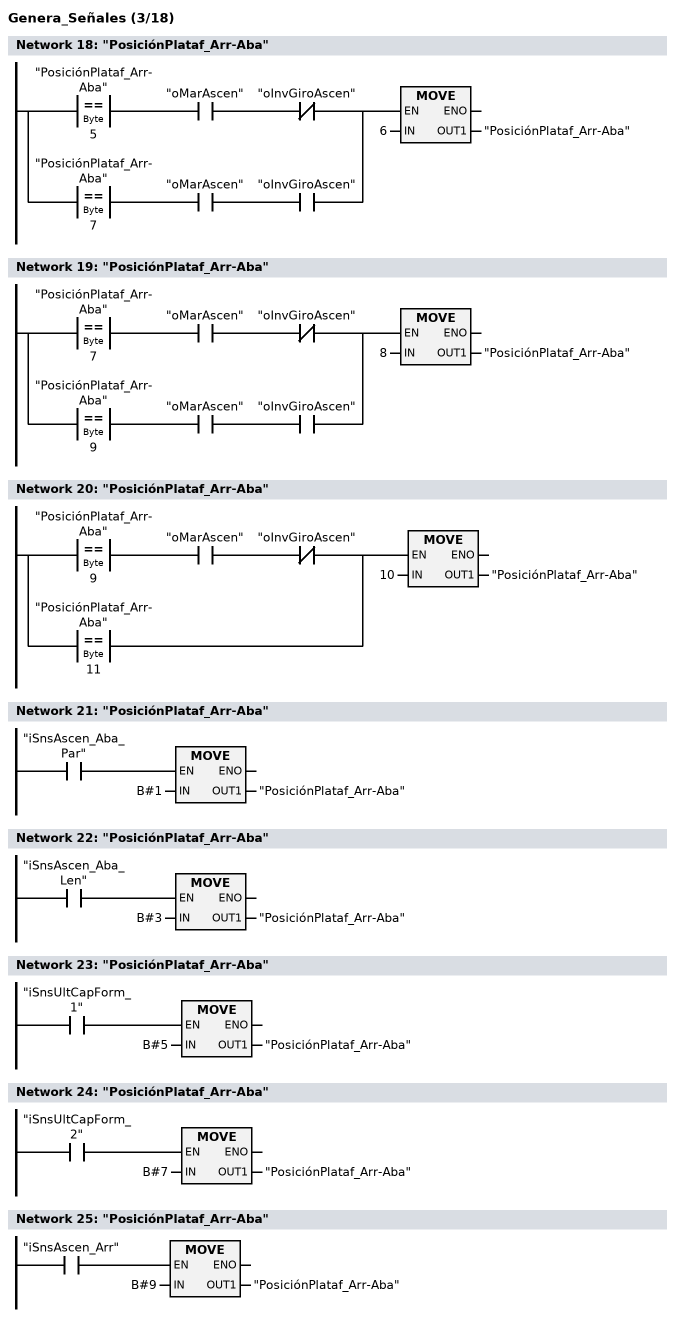
   RUNG wire#powerrail
      { S7_Templates := "SrcType := Byte" } EQ_Contact(in1 := "PosiciónPlataf_Arr-Aba", in2 := 5)
      Contact( "oMarAscen" )
      I_Contact( "oInvGiroAscen" )
      wire#w1
      { S7_GenerateENO := "TRUE" } Move(in := 6, out1 => "PosiciónPlataf_Arr-Aba")
   END_RUNG
   RUNG wire#powerrail
      { S7_Templates := "SrcType := Byte" } EQ_Contact(in1 := "PosiciónPlataf_Arr-Aba", in2 := 7)
      Contact( "oMarAscen" )
      Contact( "oInvGiroAscen" )
   END_RUNG wire#w1
   // the same network as SCL:
   IF (("PosiciónPlataf_Arr-Aba" = 5) AND "oMarAscen" AND NOT "oInvGiroAscen") OR (("PosiciónPlataf_Arr-Aba" = 7) AND "oMarAscen" AND "oInvGiroAscen") THEN
       "PosiciónPlataf_Arr-Aba" := 6;
   END_IF;
END_REGION

REGION Network 19: "PosiciónPlataf_Arr-Aba"
   RUNG wire#powerrail
      { S7_Templates := "SrcType := Byte" } EQ_Contact(in1 := "PosiciónPlataf_Arr-Aba", in2 := 7)
      Contact( "oMarAscen" )
      I_Contact( "oInvGiroAscen" )
      wire#w1
      { S7_GenerateENO := "TRUE" } Move(in := 8, out1 => "PosiciónPlataf_Arr-Aba")
   END_RUNG
   RUNG wire#powerrail
      { S7_Templates := "SrcType := Byte" } EQ_Contact(in1 := "PosiciónPlataf_Arr-Aba", in2 := 9)
      Contact( "oMarAscen" )
      Contact( "oInvGiroAscen" )
   END_RUNG wire#w1
   // the same network as SCL:
   IF (("PosiciónPlataf_Arr-Aba" = 7) AND "oMarAscen" AND NOT "oInvGiroAscen") OR (("PosiciónPlataf_Arr-Aba" = 9) AND "oMarAscen" AND "oInvGiroAscen") THEN
       "PosiciónPlataf_Arr-Aba" := 8;
   END_IF;
END_REGION

REGION Network 20: "PosiciónPlataf_Arr-Aba"
   RUNG wire#powerrail
      { S7_Templates := "SrcType := Byte" } EQ_Contact(in1 := "PosiciónPlataf_Arr-Aba", in2 := 9)
      Contact( "oMarAscen" )
      I_Contact( "oInvGiroAscen" )
      wire#w1
      { S7_GenerateENO := "TRUE" } Move(in := 10, out1 => "PosiciónPlataf_Arr-Aba")
   END_RUNG
   RUNG wire#powerrail
      { S7_Templates := "SrcType := Byte" } EQ_Contact(in1 := "PosiciónPlataf_Arr-Aba", in2 := 11)
   END_RUNG wire#w1
   // the same network as SCL:
   IF (("PosiciónPlataf_Arr-Aba" = 9) AND "oMarAscen" AND NOT "oInvGiroAscen") OR ("PosiciónPlataf_Arr-Aba" = 11) THEN
       "PosiciónPlataf_Arr-Aba" := 10;
   END_IF;
END_REGION

REGION Network 21: "PosiciónPlataf_Arr-Aba"
   RUNG wire#powerrail
      Contact( "iSnsAscen_Aba_Par" )
      { S7_GenerateENO := "TRUE" } Move(in := B#1, out1 => "PosiciónPlataf_Arr-Aba")
   END_RUNG
   // the same network as SCL:
   IF "iSnsAscen_Aba_Par" THEN "PosiciónPlataf_Arr-Aba" := B#1; END_IF;
END_REGION

REGION Network 22: "PosiciónPlataf_Arr-Aba"
   RUNG wire#powerrail
      Contact( "iSnsAscen_Aba_Len" )
      { S7_GenerateENO := "TRUE" } Move(in := B#3, out1 => "PosiciónPlataf_Arr-Aba")
   END_RUNG
   // the same network as SCL:
   IF "iSnsAscen_Aba_Len" THEN "PosiciónPlataf_Arr-Aba" := B#3; END_IF;
END_REGION

REGION Network 23: "PosiciónPlataf_Arr-Aba"
   RUNG wire#powerrail
      Contact( "iSnsUltCapForm_1" )
      { S7_GenerateENO := "TRUE" } Move(in := B#5, out1 => "PosiciónPlataf_Arr-Aba")
   END_RUNG
   // the same network as SCL:
   IF "iSnsUltCapForm_1" THEN "PosiciónPlataf_Arr-Aba" := B#5; END_IF;
END_REGION

REGION Network 24: "PosiciónPlataf_Arr-Aba"
   RUNG wire#powerrail
      Contact( "iSnsUltCapForm_2" )
      { S7_GenerateENO := "TRUE" } Move(in := B#7, out1 => "PosiciónPlataf_Arr-Aba")
   END_RUNG
   // the same network as SCL:
   IF "iSnsUltCapForm_2" THEN "PosiciónPlataf_Arr-Aba" := B#7; END_IF;
END_REGION

REGION Network 25: "PosiciónPlataf_Arr-Aba"
   RUNG wire#powerrail
      Contact( "iSnsAscen_Arr" )
      { S7_GenerateENO := "TRUE" } Move(in := B#9, out1 => "PosiciónPlataf_Arr-Aba")
   END_RUNG
   // the same network as SCL:
   IF "iSnsAscen_Arr" THEN "PosiciónPlataf_Arr-Aba" := B#9; END_IF;
END_REGION

REGION Network 26: "PosiciónPlataf_Arr-Aba"
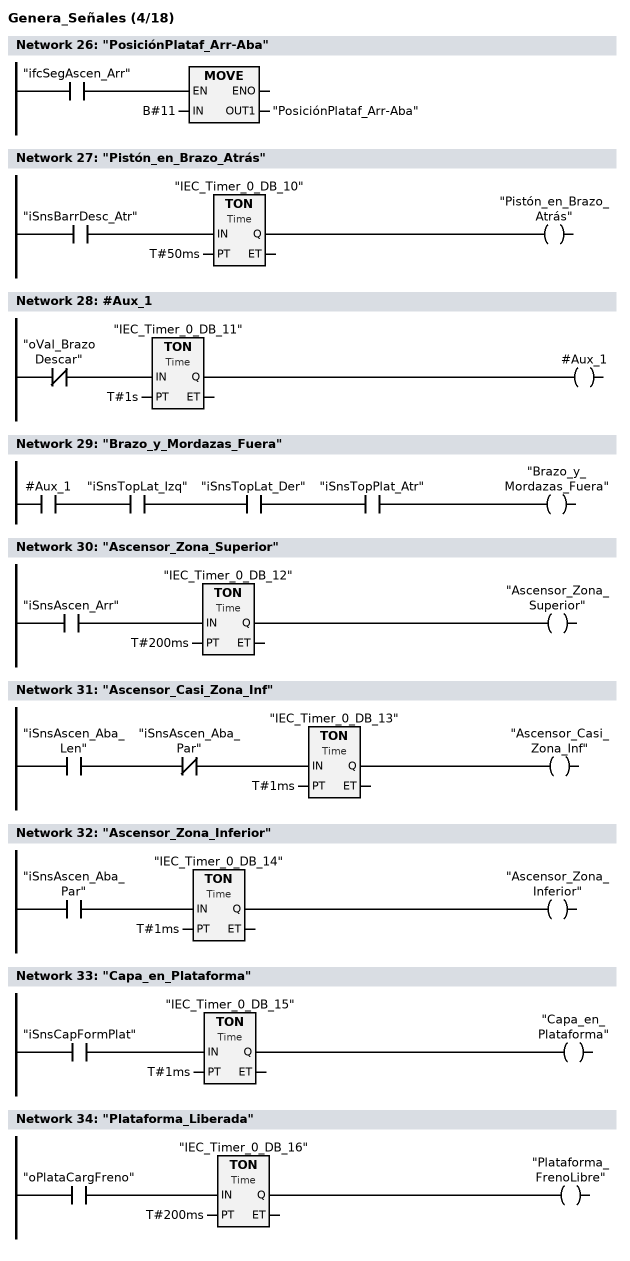
   RUNG wire#powerrail
      Contact( "ifcSegAscen_Arr" )
      { S7_GenerateENO := "TRUE" } Move(in := B#11, out1 => "PosiciónPlataf_Arr-Aba")
   END_RUNG
   // the same network as SCL:
   IF "ifcSegAscen_Arr" THEN "PosiciónPlataf_Arr-Aba" := B#11; END_IF;
END_REGION

REGION Network 27: "Pistón_en_Brazo_Atrás"
   "IEC_Timer_0_DB_10".TON(IN := "iSnsBarrDesc_Atr", PT := T#50ms);
   "Pistón_en_Brazo_Atrás" := "IEC_Timer_0_DB_10".Q;
END_REGION

REGION Network 28: #Aux_1
   "IEC_Timer_0_DB_11".TON(IN := NOT "oVal_BrazoDescar", PT := T#1s);
   #Aux_1 := "IEC_Timer_0_DB_11".Q;
END_REGION

REGION Network 29: "Brazo_y_Mordazas_Fuera"
   RUNG wire#powerrail
      Contact( #Aux_1 )
      Contact( "iSnsTopLat_Izq" )
      Contact( "iSnsTopLat_Der" )
      Contact( "iSnsTopPlat_Atr" )
      Coil( "Brazo_y_Mordazas_Fuera" )
   END_RUNG
   // the same network as SCL:
   "Brazo_y_Mordazas_Fuera" := #Aux_1 AND "iSnsTopLat_Izq" AND "iSnsTopLat_Der" AND "iSnsTopPlat_Atr";
END_REGION

REGION Network 30: "Ascensor_Zona_Superior"
   "IEC_Timer_0_DB_12".TON(IN := "iSnsAscen_Arr", PT := T#200ms);
   "Ascensor_Zona_Superior" := "IEC_Timer_0_DB_12".Q;
END_REGION

REGION Network 31: "Ascensor_Casi_Zona_Inf"
   "IEC_Timer_0_DB_13".TON(IN := "iSnsAscen_Aba_Len" AND NOT "iSnsAscen_Aba_Par", PT := T#1ms);
   "Ascensor_Casi_Zona_Inf" := "IEC_Timer_0_DB_13".Q;
END_REGION

REGION Network 32: "Ascensor_Zona_Inferior"
   "IEC_Timer_0_DB_14".TON(IN := "iSnsAscen_Aba_Par", PT := T#1ms);
   "Ascensor_Zona_Inferior" := "IEC_Timer_0_DB_14".Q;
END_REGION

REGION Network 33: "Capa_en_Plataforma"
   "IEC_Timer_0_DB_15".TON(IN := "iSnsCapFormPlat", PT := T#1ms);
   "Capa_en_Plataforma" := "IEC_Timer_0_DB_15".Q;
END_REGION

REGION Network 34: "Plataforma_Liberada"
   "IEC_Timer_0_DB_16".TON(IN := "oPlataCargFreno", PT := T#200ms);
   "Plataforma_FrenoLibre" := "IEC_Timer_0_DB_16".Q;
END_REGION

REGION Network 35: "Última_Capa" en Conteo_AUTO
END_REGION

REGION Network 36: "Brazo_Descarga_Man"
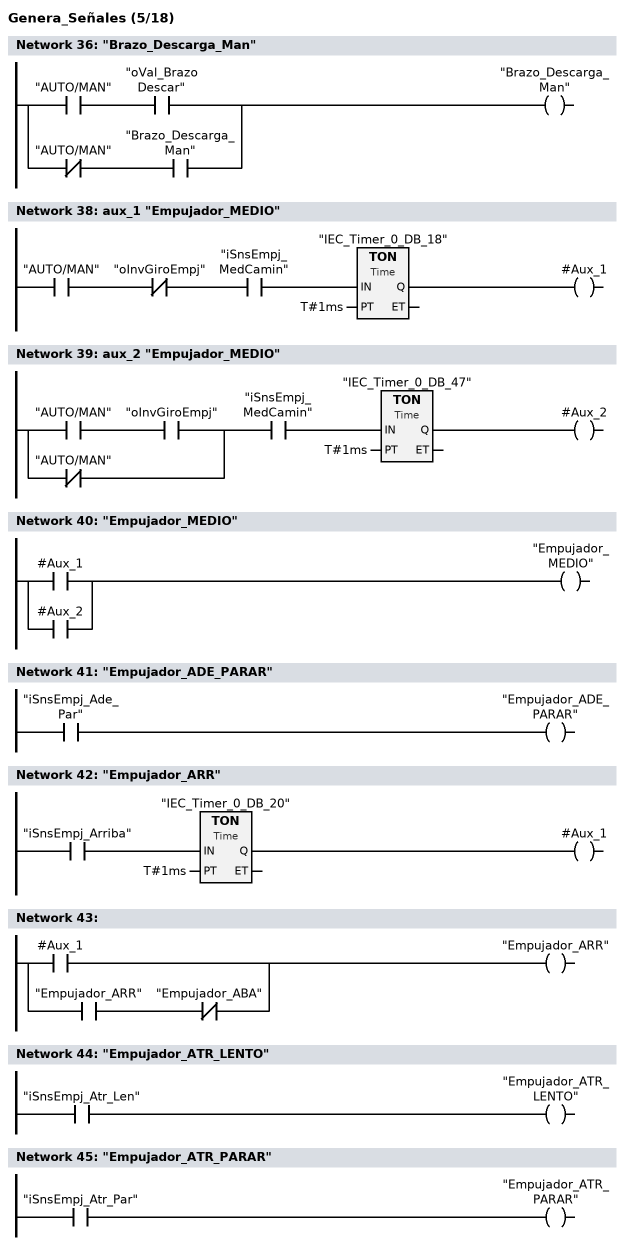
   RUNG wire#powerrail
      Contact( "AUTO/MAN" )
      Contact( "oVal_BrazoDescar" )
      wire#w1
      Coil( "Brazo_Descarga_Man" )
   END_RUNG
   RUNG wire#powerrail
      I_Contact( "AUTO/MAN" )
      Contact( "Brazo_Descarga_Man" )
   END_RUNG wire#w1
   // the same network as SCL:
   "Brazo_Descarga_Man" := ("AUTO/MAN" AND "oVal_BrazoDescar") OR (NOT "AUTO/MAN" AND "Brazo_Descarga_Man");
END_REGION

REGION Network 37: ----------------------------------------------------------------- EMPUJADOR -----------------------------------------------------------------¬
END_REGION

REGION Network 38: aux_1 "Empujador_MEDIO"
   "IEC_Timer_0_DB_18".TON(IN := "AUTO/MAN" AND NOT "oInvGiroEmpj" AND "iSnsEmpj_MedCamin", PT := T#1ms);
   #Aux_1 := "IEC_Timer_0_DB_18".Q;
END_REGION

REGION Network 39: aux_2 "Empujador_MEDIO"
   "IEC_Timer_0_DB_47".TON(IN := (("AUTO/MAN" AND "oInvGiroEmpj") OR NOT "AUTO/MAN") AND "iSnsEmpj_MedCamin",
                           PT := T#1ms);
   #Aux_2 := "IEC_Timer_0_DB_47".Q;
END_REGION

REGION Network 40: "Empujador_MEDIO"
   RUNG wire#powerrail
      Contact( #Aux_1 )
      wire#w1
      Coil( "Empujador_MEDIO" )
   END_RUNG
   RUNG wire#powerrail
      Contact( #Aux_2 )
   END_RUNG wire#w1
   // the same network as SCL:
   "Empujador_MEDIO" := #Aux_1 OR #Aux_2;
END_REGION

REGION Network 41: "Empujador_ADE_PARAR"
   RUNG wire#powerrail
      Contact( "iSnsEmpj_Ade_Par" )
      Coil( "Empujador_ADE_PARAR" )
   END_RUNG
   // the same network as SCL:
   "Empujador_ADE_PARAR" := "iSnsEmpj_Ade_Par";
END_REGION

REGION Network 42: "Empujador_ARR"
   "IEC_Timer_0_DB_20".TON(IN := "iSnsEmpj_Arriba", PT := T#1ms);
   #Aux_1 := "IEC_Timer_0_DB_20".Q;
END_REGION

REGION Network 43
   RUNG wire#powerrail
      Contact( #Aux_1 )
      wire#w1
      Coil( "Empujador_ARR" )
   END_RUNG
   RUNG wire#powerrail
      Contact( "Empujador_ARR" )
      I_Contact( "Empujador_ABA" )
   END_RUNG wire#w1
   // the same network as SCL:
   "Empujador_ARR" := #Aux_1 OR ("Empujador_ARR" AND NOT "Empujador_ABA");
END_REGION

REGION Network 44: "Empujador_ATR_LENTO"
   RUNG wire#powerrail
      Contact( "iSnsEmpj_Atr_Len" )
      Coil( "Empujador_ATR_LENTO" )
   END_RUNG
   // the same network as SCL:
   "Empujador_ATR_LENTO" := "iSnsEmpj_Atr_Len";
END_REGION

REGION Network 45: "Empujador_ATR_PARAR"
   RUNG wire#powerrail
      Contact( "iSnsEmpj_Atr_Par" )
      Coil( "Empujador_ATR_PARAR" )
   END_RUNG
   // the same network as SCL:
   "Empujador_ATR_PARAR" := "iSnsEmpj_Atr_Par";
END_REGION

REGION Network 46: "Empujador_ADE_LENTO"
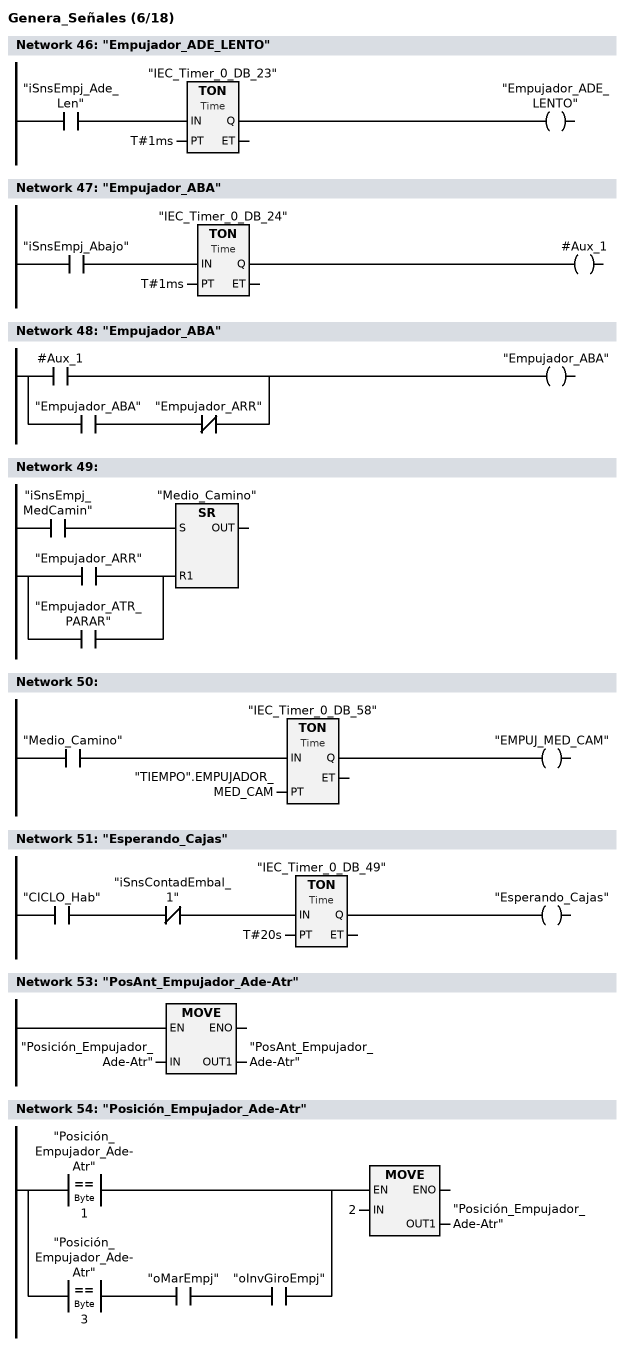
   "IEC_Timer_0_DB_23".TON(IN := "iSnsEmpj_Ade_Len", PT := T#1ms);
   "Empujador_ADE_LENTO" := "IEC_Timer_0_DB_23".Q;
END_REGION

REGION Network 47: "Empujador_ABA"
   "IEC_Timer_0_DB_24".TON(IN := "iSnsEmpj_Abajo", PT := T#1ms);
   #Aux_1 := "IEC_Timer_0_DB_24".Q;
END_REGION

REGION Network 48: "Empujador_ABA"
   RUNG wire#powerrail
      Contact( #Aux_1 )
      wire#w1
      Coil( "Empujador_ABA" )
   END_RUNG
   RUNG wire#powerrail
      Contact( "Empujador_ABA" )
      I_Contact( "Empujador_ARR" )
   END_RUNG wire#w1
   // the same network as SCL:
   "Empujador_ABA" := #Aux_1 OR ("Empujador_ABA" AND NOT "Empujador_ARR");
END_REGION

REGION Network 49
   RUNG wire#powerrail
      Contact( "iSnsEmpj_MedCamin" )
      S_SR(operand := "Medio_Camino", r1 := wire#w1)
   END_RUNG
   RUNG wire#powerrail
      Contact( "Empujador_ARR" )
   END_RUNG wire#w1
   RUNG wire#powerrail
      Contact( "Empujador_ATR_PARAR" )
   END_RUNG wire#w1
   // the same network as SCL:
   IF "iSnsEmpj_MedCamin" THEN
       "Medio_Camino" := TRUE;   // SR flip-flop
   END_IF;
   IF "Empujador_ARR" OR "Empujador_ATR_PARAR" THEN "Medio_Camino" := FALSE; END_IF;
END_REGION

REGION Network 50
   "IEC_Timer_0_DB_58".TON(IN := "Medio_Camino", PT := "TIEMPO".EMPUJADOR_MED_CAM);
   "EMPUJ_MED_CAM" := "IEC_Timer_0_DB_58".Q;
END_REGION

REGION Network 51: "Esperando_Cajas"
   "IEC_Timer_0_DB_49".TON(IN := "CICLO_Hab" AND NOT "iSnsContadEmbal_1", PT := T#20s);
   "Esperando_Cajas" := "IEC_Timer_0_DB_49".Q;
END_REGION

REGION Network 52: ------------------------------------------------------------------------------------------------------------------------------------------------------------
END_REGION

REGION Network 53: "PosAnt_Empujador_Ade-Atr"
   RUNG wire#powerrail
      { S7_GenerateENO := "TRUE" } Move(in := "Posición_Empujador_Ade-Atr", out1 => "PosAnt_Empujador_Ade-Atr")
   END_RUNG
   // the same network as SCL:
   "PosAnt_Empujador_Ade-Atr" := "Posición_Empujador_Ade-Atr";
END_REGION

REGION Network 54: "Posición_Empujador_Ade-Atr"
   RUNG wire#powerrail
      { S7_Templates := "SrcType := Byte" } EQ_Contact(in1 := "Posición_Empujador_Ade-Atr", in2 := 1)
      wire#w1
      { S7_GenerateENO := "TRUE" } Move(in := 2, out1 => "Posición_Empujador_Ade-Atr")
   END_RUNG
   RUNG wire#powerrail
      { S7_Templates := "SrcType := Byte" } EQ_Contact(in1 := "Posición_Empujador_Ade-Atr", in2 := 3)
      Contact( "oMarEmpj" )
      Contact( "oInvGiroEmpj" )
   END_RUNG wire#w1
   // the same network as SCL:
   IF ("Posición_Empujador_Ade-Atr" = 1) OR (("Posición_Empujador_Ade-Atr" = 3) AND "oMarEmpj" AND "oInvGiroEmpj") THEN
       "Posición_Empujador_Ade-Atr" := 2;
   END_IF;
END_REGION

REGION Network 55: "Posición_Empujador_Ade-Atr"
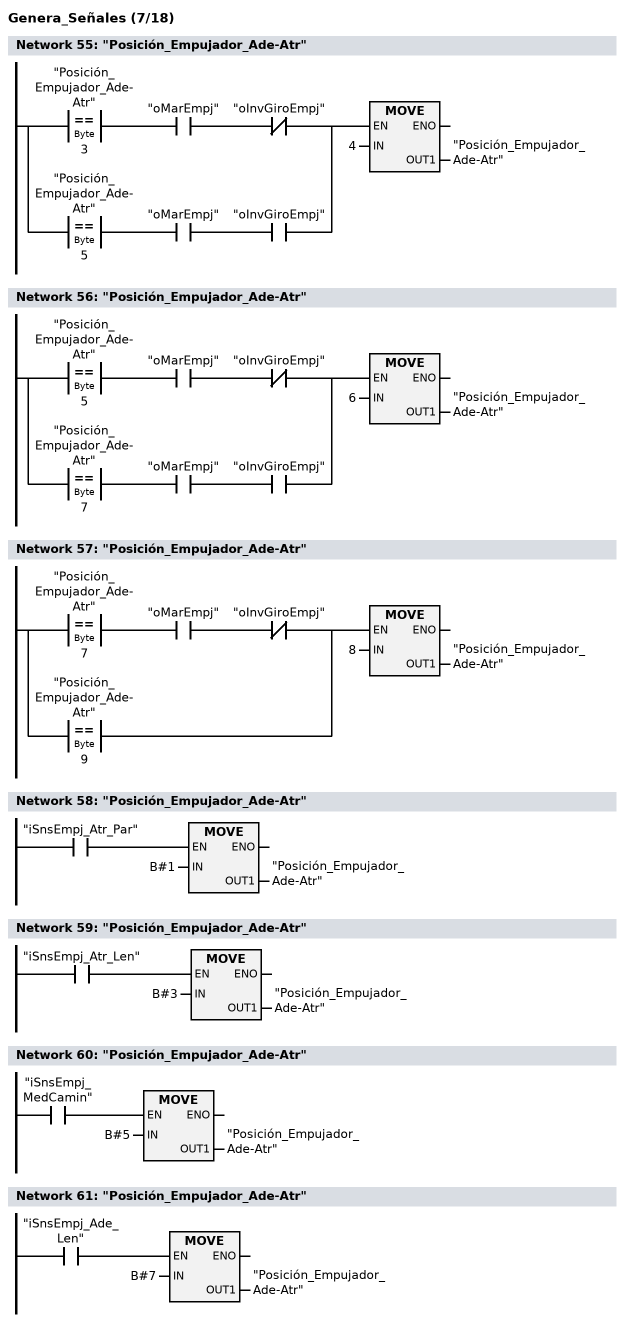
   RUNG wire#powerrail
      { S7_Templates := "SrcType := Byte" } EQ_Contact(in1 := "Posición_Empujador_Ade-Atr", in2 := 3)
      Contact( "oMarEmpj" )
      I_Contact( "oInvGiroEmpj" )
      wire#w1
      { S7_GenerateENO := "TRUE" } Move(in := 4, out1 => "Posición_Empujador_Ade-Atr")
   END_RUNG
   RUNG wire#powerrail
      { S7_Templates := "SrcType := Byte" } EQ_Contact(in1 := "Posición_Empujador_Ade-Atr", in2 := 5)
      Contact( "oMarEmpj" )
      Contact( "oInvGiroEmpj" )
   END_RUNG wire#w1
   // the same network as SCL:
   IF (("Posición_Empujador_Ade-Atr" = 3) AND "oMarEmpj" AND NOT "oInvGiroEmpj") OR (("Posición_Empujador_Ade-Atr" = 5) AND "oMarEmpj" AND "oInvGiroEmpj") THEN
       "Posición_Empujador_Ade-Atr" := 4;
   END_IF;
END_REGION

REGION Network 56: "Posición_Empujador_Ade-Atr"
   RUNG wire#powerrail
      { S7_Templates := "SrcType := Byte" } EQ_Contact(in1 := "Posición_Empujador_Ade-Atr", in2 := 5)
      Contact( "oMarEmpj" )
      I_Contact( "oInvGiroEmpj" )
      wire#w1
      { S7_GenerateENO := "TRUE" } Move(in := 6, out1 => "Posición_Empujador_Ade-Atr")
   END_RUNG
   RUNG wire#powerrail
      { S7_Templates := "SrcType := Byte" } EQ_Contact(in1 := "Posición_Empujador_Ade-Atr", in2 := 7)
      Contact( "oMarEmpj" )
      Contact( "oInvGiroEmpj" )
   END_RUNG wire#w1
   // the same network as SCL:
   IF (("Posición_Empujador_Ade-Atr" = 5) AND "oMarEmpj" AND NOT "oInvGiroEmpj") OR (("Posición_Empujador_Ade-Atr" = 7) AND "oMarEmpj" AND "oInvGiroEmpj") THEN
       "Posición_Empujador_Ade-Atr" := 6;
   END_IF;
END_REGION

REGION Network 57: "Posición_Empujador_Ade-Atr"
   RUNG wire#powerrail
      { S7_Templates := "SrcType := Byte" } EQ_Contact(in1 := "Posición_Empujador_Ade-Atr", in2 := 7)
      Contact( "oMarEmpj" )
      I_Contact( "oInvGiroEmpj" )
      wire#w1
      { S7_GenerateENO := "TRUE" } Move(in := 8, out1 => "Posición_Empujador_Ade-Atr")
   END_RUNG
   RUNG wire#powerrail
      { S7_Templates := "SrcType := Byte" } EQ_Contact(in1 := "Posición_Empujador_Ade-Atr", in2 := 9)
   END_RUNG wire#w1
   // the same network as SCL:
   IF (("Posición_Empujador_Ade-Atr" = 7) AND "oMarEmpj" AND NOT "oInvGiroEmpj") OR ("Posición_Empujador_Ade-Atr" = 9) THEN
       "Posición_Empujador_Ade-Atr" := 8;
   END_IF;
END_REGION

REGION Network 58: "Posición_Empujador_Ade-Atr"
   RUNG wire#powerrail
      Contact( "iSnsEmpj_Atr_Par" )
      { S7_GenerateENO := "TRUE" } Move(in := B#1, out1 => "Posición_Empujador_Ade-Atr")
   END_RUNG
   // the same network as SCL:
   IF "iSnsEmpj_Atr_Par" THEN "Posición_Empujador_Ade-Atr" := B#1; END_IF;
END_REGION

REGION Network 59: "Posición_Empujador_Ade-Atr"
   RUNG wire#powerrail
      Contact( "iSnsEmpj_Atr_Len" )
      { S7_GenerateENO := "TRUE" } Move(in := B#3, out1 => "Posición_Empujador_Ade-Atr")
   END_RUNG
   // the same network as SCL:
   IF "iSnsEmpj_Atr_Len" THEN "Posición_Empujador_Ade-Atr" := B#3; END_IF;
END_REGION

REGION Network 60: "Posición_Empujador_Ade-Atr"
   RUNG wire#powerrail
      Contact( "iSnsEmpj_MedCamin" )
      { S7_GenerateENO := "TRUE" } Move(in := B#5, out1 => "Posición_Empujador_Ade-Atr")
   END_RUNG
   // the same network as SCL:
   IF "iSnsEmpj_MedCamin" THEN "Posición_Empujador_Ade-Atr" := B#5; END_IF;
END_REGION

REGION Network 61: "Posición_Empujador_Ade-Atr"
   RUNG wire#powerrail
      Contact( "iSnsEmpj_Ade_Len" )
      { S7_GenerateENO := "TRUE" } Move(in := B#7, out1 => "Posición_Empujador_Ade-Atr")
   END_RUNG
   // the same network as SCL:
   IF "iSnsEmpj_Ade_Len" THEN "Posición_Empujador_Ade-Atr" := B#7; END_IF;
END_REGION

REGION Network 62: "Posición_Empujador_Ade-Atr"
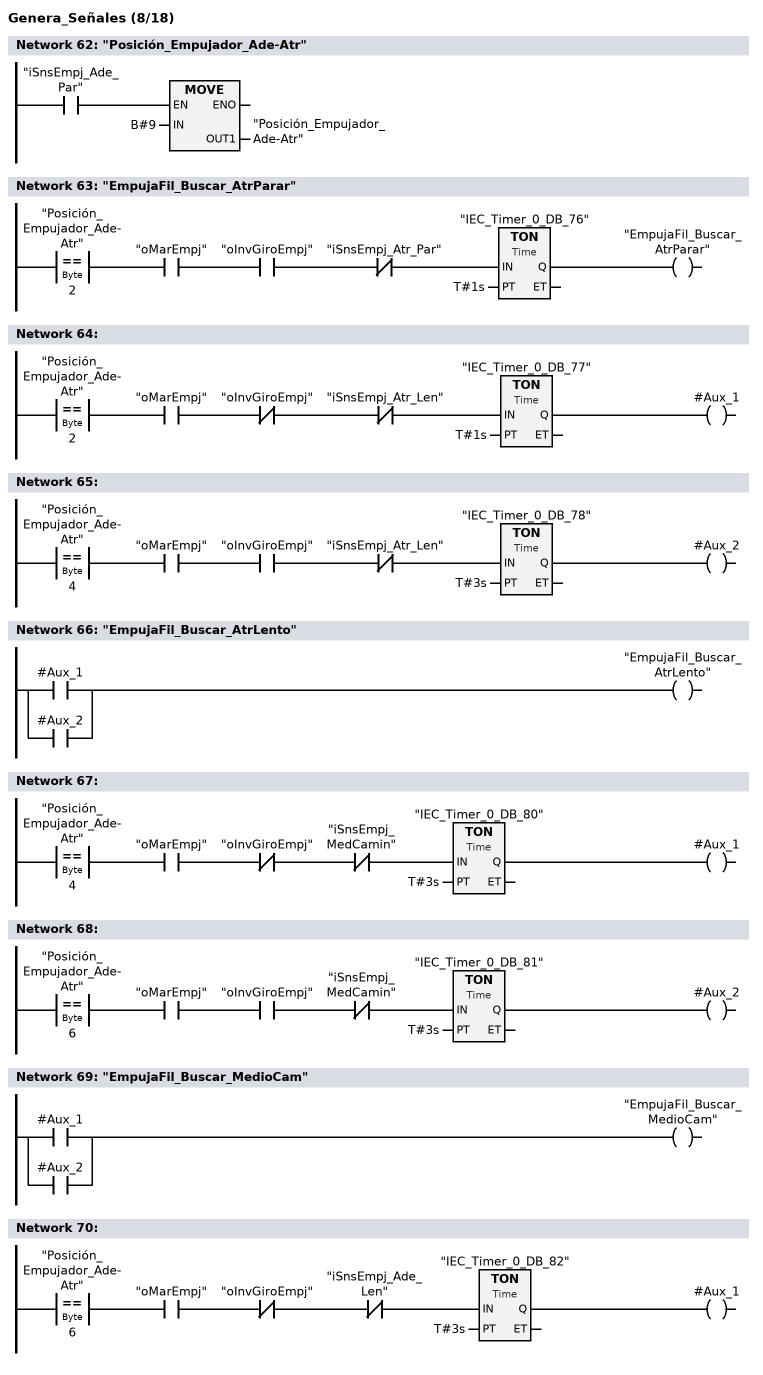
   RUNG wire#powerrail
      Contact( "iSnsEmpj_Ade_Par" )
      { S7_GenerateENO := "TRUE" } Move(in := B#9, out1 => "Posición_Empujador_Ade-Atr")
   END_RUNG
   // the same network as SCL:
   IF "iSnsEmpj_Ade_Par" THEN "Posición_Empujador_Ade-Atr" := B#9; END_IF;
END_REGION

REGION Network 63: "EmpujaFil_Buscar_AtrParar"
   "IEC_Timer_0_DB_76".TON(IN := ("Posición_Empujador_Ade-Atr" = 2) AND "oMarEmpj" AND "oInvGiroEmpj" AND NOT "iSnsEmpj_Atr_Par",
                           PT := T#1s);
   "EmpujaFil_Buscar_AtrParar" := "IEC_Timer_0_DB_76".Q;
END_REGION

REGION Network 64
   "IEC_Timer_0_DB_77".TON(IN := ("Posición_Empujador_Ade-Atr" = 2) AND "oMarEmpj" AND NOT "oInvGiroEmpj" AND NOT "iSnsEmpj_Atr_Len",
                           PT := T#1s);
   #Aux_1 := "IEC_Timer_0_DB_77".Q;
END_REGION

REGION Network 65
   "IEC_Timer_0_DB_78".TON(IN := ("Posición_Empujador_Ade-Atr" = 4) AND "oMarEmpj" AND "oInvGiroEmpj" AND NOT "iSnsEmpj_Atr_Len",
                           PT := T#3s);
   #Aux_2 := "IEC_Timer_0_DB_78".Q;
END_REGION

REGION Network 66: "EmpujaFil_Buscar_AtrLento"
   RUNG wire#powerrail
      Contact( #Aux_1 )
      wire#w1
      Coil( "EmpujaFil_Buscar_AtrLento" )
   END_RUNG
   RUNG wire#powerrail
      Contact( #Aux_2 )
   END_RUNG wire#w1
   // the same network as SCL:
   "EmpujaFil_Buscar_AtrLento" := #Aux_1 OR #Aux_2;
END_REGION

REGION Network 67
   "IEC_Timer_0_DB_80".TON(IN := ("Posición_Empujador_Ade-Atr" = 4) AND "oMarEmpj" AND NOT "oInvGiroEmpj" AND NOT "iSnsEmpj_MedCamin",
                           PT := T#3s);
   #Aux_1 := "IEC_Timer_0_DB_80".Q;
END_REGION

REGION Network 68
   "IEC_Timer_0_DB_81".TON(IN := ("Posición_Empujador_Ade-Atr" = 6) AND "oMarEmpj" AND "oInvGiroEmpj" AND NOT "iSnsEmpj_MedCamin",
                           PT := T#3s);
   #Aux_2 := "IEC_Timer_0_DB_81".Q;
END_REGION

REGION Network 69: "EmpujaFil_Buscar_MedioCam"
   RUNG wire#powerrail
      Contact( #Aux_1 )
      wire#w1
      Coil( "EmpujaFil_Buscar_MedioCam" )
   END_RUNG
   RUNG wire#powerrail
      Contact( #Aux_2 )
   END_RUNG wire#w1
   // the same network as SCL:
   "EmpujaFil_Buscar_MedioCam" := #Aux_1 OR #Aux_2;
END_REGION

REGION Network 70
   "IEC_Timer_0_DB_82".TON(IN := ("Posición_Empujador_Ade-Atr" = 6) AND "oMarEmpj" AND NOT "oInvGiroEmpj" AND NOT "iSnsEmpj_Ade_Len",
                           PT := T#3s);
   #Aux_1 := "IEC_Timer_0_DB_82".Q;
END_REGION

REGION Network 71
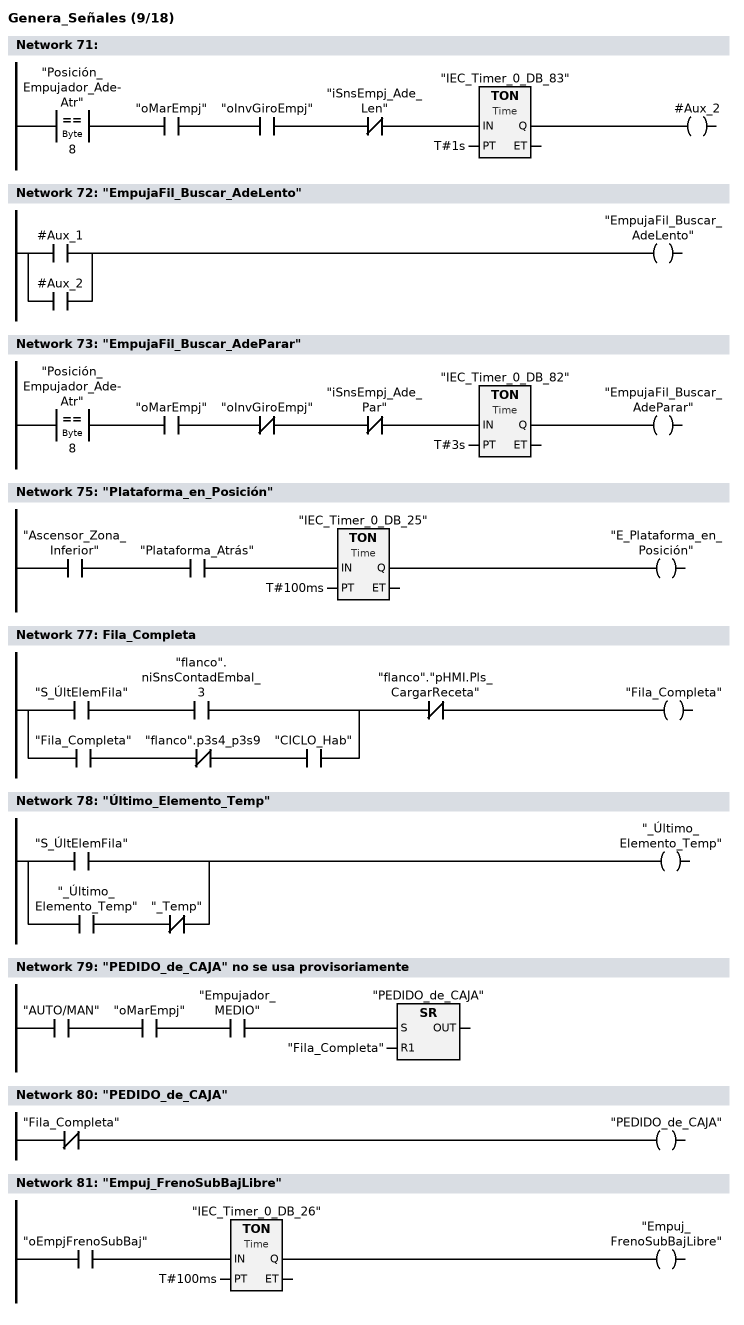
   "IEC_Timer_0_DB_83".TON(IN := ("Posición_Empujador_Ade-Atr" = 8) AND "oMarEmpj" AND "oInvGiroEmpj" AND NOT "iSnsEmpj_Ade_Len",
                           PT := T#1s);
   #Aux_2 := "IEC_Timer_0_DB_83".Q;
END_REGION

REGION Network 72: "EmpujaFil_Buscar_AdeLento"
   RUNG wire#powerrail
      Contact( #Aux_1 )
      wire#w1
      Coil( "EmpujaFil_Buscar_AdeLento" )
   END_RUNG
   RUNG wire#powerrail
      Contact( #Aux_2 )
   END_RUNG wire#w1
   // the same network as SCL:
   "EmpujaFil_Buscar_AdeLento" := #Aux_1 OR #Aux_2;
END_REGION

REGION Network 73: "EmpujaFil_Buscar_AdeParar"
   "IEC_Timer_0_DB_82".TON(IN := ("Posición_Empujador_Ade-Atr" = 8) AND "oMarEmpj" AND NOT "oInvGiroEmpj" AND NOT "iSnsEmpj_Ade_Par",
                           PT := T#3s);
   "EmpujaFil_Buscar_AdeParar" := "IEC_Timer_0_DB_82".Q;
END_REGION

REGION Network 74: ---------------------------------------------------------------------------------------------------------------------------------------------------------------------------
END_REGION

REGION Network 75: "Plataforma_en_Posición"
   "IEC_Timer_0_DB_25".TON(IN := "Ascensor_Zona_Inferior" AND "Plataforma_Atrás", PT := T#100ms);
   "E_Plataforma_en_Posición" := "IEC_Timer_0_DB_25".Q;
END_REGION

REGION Network 77: Fila_Completa
   RUNG wire#powerrail
      Contact( "S_ÚltElemFila" )
      Contact( "flanco".niSnsContadEmbal_3 )
      wire#w1
      I_Contact( "flanco"."pHMI.Pls_CargarReceta" )
      Coil( "Fila_Completa" )
   END_RUNG
   RUNG wire#powerrail
      Contact( "Fila_Completa" )
      I_Contact( "flanco".p3s4_p3s9 )
      Contact( "CICLO_Hab" )
   END_RUNG wire#w1
   // the same network as SCL:
   "Fila_Completa" := (("S_ÚltElemFila" AND "flanco".niSnsContadEmbal_3) OR ("Fila_Completa" AND NOT "flanco".p3s4_p3s9 AND "CICLO_Hab")) AND NOT "flanco"."pHMI.Pls_CargarReceta";
END_REGION

REGION Network 78: "Último_Elemento_Temp"
   RUNG wire#powerrail
      Contact( "S_ÚltElemFila" )
      wire#w1
      Coil( "_Último_Elemento_Temp" )
   END_RUNG
   RUNG wire#powerrail
      Contact( "_Último_Elemento_Temp" )
      I_Contact( "_Temp" )
   END_RUNG wire#w1
   // the same network as SCL:
   "_Último_Elemento_Temp" := "S_ÚltElemFila" OR ("_Último_Elemento_Temp" AND NOT "_Temp");
END_REGION

REGION Network 79: "PEDIDO_de_CAJA" no se usa provisoriamente
   RUNG wire#powerrail
      Contact( "AUTO/MAN" )
      Contact( "oMarEmpj" )
      Contact( "Empujador_MEDIO" )
      S_SR(operand := "PEDIDO_de_CAJA", r1 := "Fila_Completa")
   END_RUNG
   // the same network as SCL:
   IF "AUTO/MAN" AND "oMarEmpj" AND "Empujador_MEDIO" THEN
       "PEDIDO_de_CAJA" := TRUE;   // SR flip-flop
   END_IF;
   IF "Fila_Completa" THEN "PEDIDO_de_CAJA" := FALSE; END_IF;
END_REGION

REGION Network 80: "PEDIDO_de_CAJA"
   RUNG wire#powerrail
      I_Contact( "Fila_Completa" )
      Coil( "PEDIDO_de_CAJA" )
   END_RUNG
   // the same network as SCL:
   "PEDIDO_de_CAJA" := NOT "Fila_Completa";
END_REGION

REGION Network 81: "Empuj_FrenoSubBajLibre"
   "IEC_Timer_0_DB_26".TON(IN := "oEmpjFrenoSubBaj", PT := T#100ms);
   "Empuj_FrenoSubBajLibre" := "IEC_Timer_0_DB_26".Q;
END_REGION

REGION Network 82: "Elemento_CARGADO"
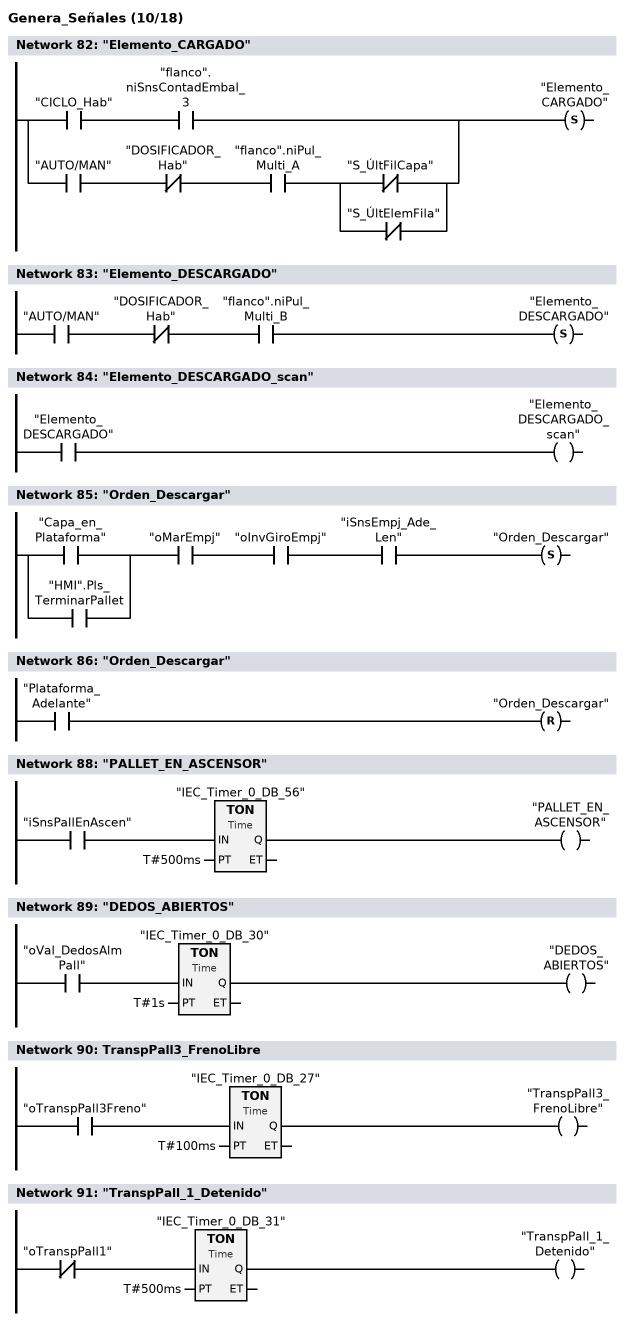
   RUNG wire#powerrail
      Contact( "CICLO_Hab" )
      Contact( "flanco".niSnsContadEmbal_3 )
      wire#w1
      S_Coil( "Elemento_CARGADO" )
   END_RUNG
   RUNG wire#powerrail
      Contact( "AUTO/MAN" )
      I_Contact( "DOSIFICADOR_Hab" )
      Contact( "flanco".niPul_Multi_A )
      wire#w2
      I_Contact( "S_ÚltFilCapa" )
   END_RUNG wire#w1
   RUNG wire#w2
      I_Contact( "S_ÚltElemFila" )
   END_RUNG wire#w1
   // the same network as SCL:
   IF ("CICLO_Hab" AND "flanco".niSnsContadEmbal_3) OR ("AUTO/MAN" AND NOT "DOSIFICADOR_Hab" AND "flanco".niPul_Multi_A AND (NOT "S_ÚltFilCapa" OR NOT "S_ÚltElemFila")) THEN
       "Elemento_CARGADO" := TRUE;
   END_IF;
END_REGION

REGION Network 83: "Elemento_DESCARGADO"
   RUNG wire#powerrail
      Contact( "AUTO/MAN" )
      I_Contact( "DOSIFICADOR_Hab" )
      Contact( "flanco".niPul_Multi_B )
      S_Coil( "Elemento_DESCARGADO" )
   END_RUNG
   // the same network as SCL:
   IF "AUTO/MAN" AND NOT "DOSIFICADOR_Hab" AND "flanco".niPul_Multi_B THEN
       "Elemento_DESCARGADO" := TRUE;
   END_IF;
END_REGION

REGION Network 84: "Elemento_DESCARGADO_scan"
   RUNG wire#powerrail
      Contact( "Elemento_DESCARGADO" )
      Coil( "Elemento_DESCARGADO_scan" )
   END_RUNG
   // the same network as SCL:
   "Elemento_DESCARGADO_scan" := "Elemento_DESCARGADO";
END_REGION

REGION Network 85: "Orden_Descargar"
   RUNG wire#powerrail
      Contact( "Capa_en_Plataforma" )
      wire#w1
      Contact( "oMarEmpj" )
      Contact( "oInvGiroEmpj" )
      Contact( "iSnsEmpj_Ade_Len" )
      S_Coil( "Orden_Descargar" )
   END_RUNG
   RUNG wire#powerrail
      Contact( "HMI".Pls_TerminarPallet )
   END_RUNG wire#w1
   // the same network as SCL:
   IF ("Capa_en_Plataforma" OR "HMI".Pls_TerminarPallet) AND "oMarEmpj" AND "oInvGiroEmpj" AND "iSnsEmpj_Ade_Len" THEN
       "Orden_Descargar" := TRUE;
   END_IF;
END_REGION

REGION Network 86: "Orden_Descargar"
   RUNG wire#powerrail
      Contact( "Plataforma_Adelante" )
      R_Coil( "Orden_Descargar" )
   END_RUNG
   // the same network as SCL:
   IF "Plataforma_Adelante" THEN "Orden_Descargar" := FALSE; END_IF;
END_REGION

REGION Network 87: ----------------------------------------------------------------- TRANSPORTE PALLETS-----------------------------------------------------------------¬
END_REGION

REGION Network 88: "PALLET_EN_ASCENSOR"
   "IEC_Timer_0_DB_56".TON(IN := "iSnsPallEnAscen", PT := T#500ms);
   "PALLET_EN_ASCENSOR" := "IEC_Timer_0_DB_56".Q;
END_REGION

REGION Network 89: "DEDOS_ABIERTOS"
   "IEC_Timer_0_DB_30".TON(IN := "oVal_DedosAlmPall", PT := T#1s);
   "DEDOS_ABIERTOS" := "IEC_Timer_0_DB_30".Q;
END_REGION

REGION Network 90: TranspPall3_FrenoLibre
   "IEC_Timer_0_DB_27".TON(IN := "oTranspPall3Freno", PT := T#100ms);
   "TranspPall3_FrenoLibre" := "IEC_Timer_0_DB_27".Q;
END_REGION

REGION Network 91: "TranspPall_1_Detenido"
   "IEC_Timer_0_DB_31".TON(IN := NOT "oTranspPall1", PT := T#500ms);
   "TranspPall_1_Detenido" := "IEC_Timer_0_DB_31".Q;
END_REGION

REGION Network 92: Aux "PALLET_EN_ASCENSOR"
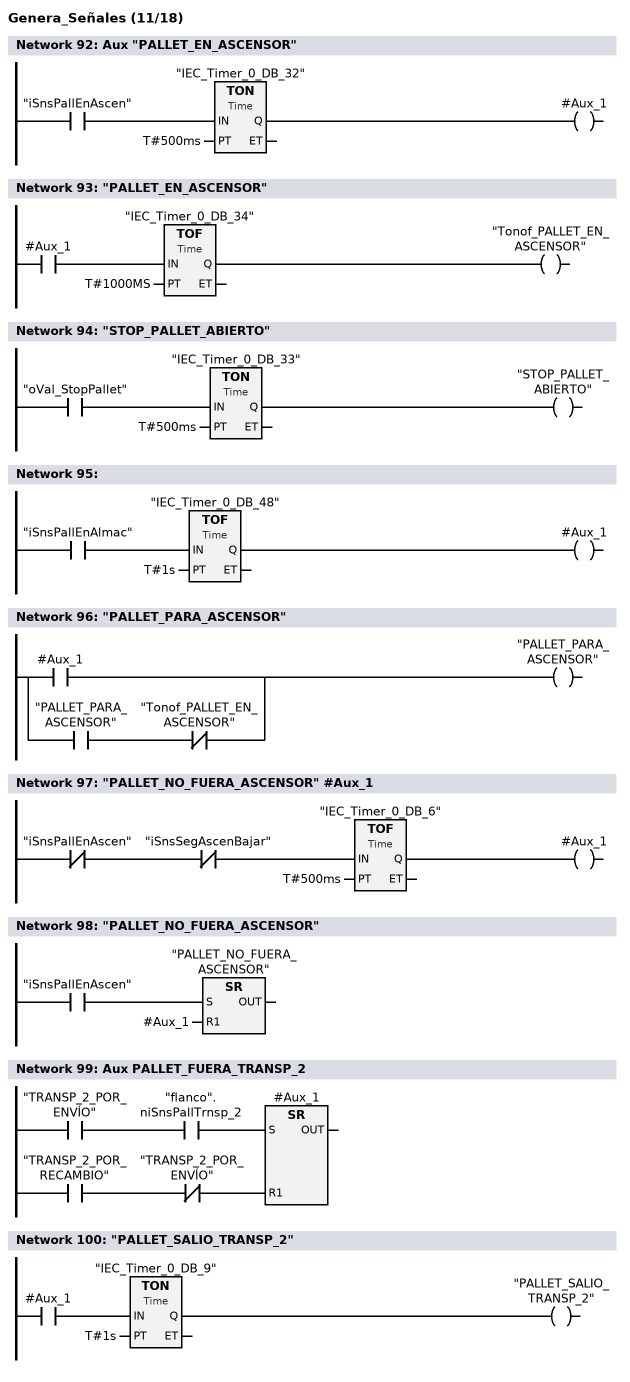
   "IEC_Timer_0_DB_32".TON(IN := "iSnsPallEnAscen", PT := T#500ms);
   #Aux_1 := "IEC_Timer_0_DB_32".Q;
END_REGION

REGION Network 93: "PALLET_EN_ASCENSOR"
   "IEC_Timer_0_DB_34".TOF(IN := #Aux_1, PT := T#1000MS);
   "Tonof_PALLET_EN_ASCENSOR" := "IEC_Timer_0_DB_34".Q;
END_REGION

REGION Network 94: "STOP_PALLET_ABIERTO"
   "IEC_Timer_0_DB_33".TON(IN := "oVal_StopPallet", PT := T#500ms);
   "STOP_PALLET_ABIERTO" := "IEC_Timer_0_DB_33".Q;
END_REGION

REGION Network 95
   "IEC_Timer_0_DB_48".TOF(IN := "iSnsPallEnAlmac", PT := T#1s);
   #Aux_1 := "IEC_Timer_0_DB_48".Q;
END_REGION
